screen "Filling" 800x480
   Button "Button_19" at 183,156 size 77x32; TextOff 'Aut'
      on Click: SetBit("Data_Tank1_Filling_Cmd_AutCtrl")
   TextField "Text field_26" at 286,75 size 190x23; Text 'Filling phase control'
   TextField "Text field_27" at 182,109 size 83x23; Text 'Automat'
   TextField "Text field_28" at 182,127 size 70x23; Text 'Manual'
   Button "Button_20" at 263,156 size 77x32; TextOff 'Man'
      on Click: SetBit("Data_Tank1_Filling_Cmd_ManCtrl")
   Circle "Circle_14" at 299,110 size 20x20
      Appearance <- "Data_Tank1_Filling_State_AutCtrl"
   Circle "Circle_15" at 299,130 size 20x20
      Appearance <- "Data_Tank1_Filling_State_ManCtrl"
   Button "Button_21" at 344,156 size 157x32; TextOff 'Reset done'
      on Click: SetBit("Data_Tank1_Filling_Cmd_ResetDone")
   Button "Button_22" at 183,206 size 77x32; TextOff 'Start'
      on Click: SetBit("Data_Tank1_Filling_Cmd_StartMan")
   Button "Button_23" at 263,205 size 77x32; TextOff 'Stop'
      on Click: SetBit("Data_Tank1_Filling_Cmd_StopMan")
   Button "Button_24" at 423,205 size 77x32; TextOff 'Rsume'
      on Click: SetBit("Data_Tank1_Filling_Cmd_ResumeMan")
   Button "Button_25" at 343,205 size 77x32; TextOff 'Pause'
      on Click: SetBit("Data_Tank1_Filling_Cmd_PauseMan")
   TextField "Text field_29" at 343,118 size 51x23; Text 'Done'
   Circle "Circle_16" at 460,119 size 20x20
      Appearance <- "Data_Tank1_Filling_State_Done"
   GraphicView "Graphic view_1" at 525,70 size 75x74; Picture "exit-png-cancel-cross-exit-remove-icon-512"
   Button "Button_26" at 520,72 size 76x81; TextOff 'Text'
      on Click: ActivateScreen("MainScr", 0)
   Group "Group" at 169,70 size 431x184; Picture "exit-png-cancel-cross-exit-remove-icon-512"
   SymbolLibrary "Symbol library_1" at 202,63 size 120x212
   SymbolLibrary "Symbol library_2" at 148,84 size 58x23
   SymbolLibrary "Symbol library_3" at 320,241 size 20x23
   Bar "Bar_1" at 204,63 size 117x211; MinimumValue 0; MaximumValue 2
      ProcessValue <- "Data_Tank1_WaterLevel_AIScaled"
   SymbolLibrary "Symbol library_4" at 55,31 size 94x80
      Appearance <- "Data_Tank1_ValveFill_State_StColor"
   IOField "I/O field_1" at 215,109 size 96x32; FormatPattern s9.99; Unit  m
      ProcessValue <- "Data_Tank1_WaterLevel_AIScaled"
   IOField "I/O field_2" at 216,143 size 96x32; FormatPattern 999.9; Unit  °C
      ProcessValue <- "Data_Tank1_WaterTemp_AIScaled"
   SymbolLibrary "Symbol library_6" at 226,190 size 71x61
      Appearance <- "Data_Tank1_Mixer_State_StateInt"
   Button "Button_1" at 7,233 size 77x32; TextOff 'Aut'
      on Click: SetBit("Data_Tank1_ValveFill_Cmd_AutCtrl")
   TextField "Text field_1" at 45,123 size 83x23; Text 'ValveFill'
   TextField "Text field_2" at 5,148 size 83x23; Text 'Automat'
   TextField "Text field_3" at 5,166 size 70x23; Text 'Manual'
   TextField "Text field_4" at 5,188 size 51x23; Text 'Open'
   TextField "Text field_5" at 5,206 size 65x23; Text 'Closed'
   Button "Button_2" at 86,233 size 77x32; TextOff 'Man'
      on Click: SetBit("Data_Tank1_ValveFill_Cmd_ManCtrl")
   Button "Button_3" at 7,267 size 77x32; TextOff 'Open'
      on Click: SetBit("Data_Tank1_ValveFill_Cmd_OpenMan")
   Button "Button_4" at 86,267 size 77x32; TextOff 'Close'
      on Click: SetBit("Data_Tank1_ValveFill_Cmd_CloseMan")
   Button "Button_5" at 419,209 size 77x32; TextOff 'Aut'
      on Click: SetBit("Data_Tank1_ValveDrain_Cmd_AutCtrl")
   TextField "Text field_6" at 450,99 size 104x23; Text 'ValveDrain'
   TextField "Text field_7" at 417,124 size 83x23; Text 'Automat'
   TextField "Text field_8" at 417,142 size 70x23; Text 'Manual'
   TextField "Text field_9" at 417,164 size 51x23; Text 'Open'
   TextField "Text field_10" at 417,182 size 65x23; Text 'Closed'
   Button "Button_6" at 498,209 size 77x32; TextOff 'Man'
      on Click: SetBit("Data_Tank1_Mixer_Cmd_ManCtrl")
   TextField "Text field_11" at 234,284 size 56x23; Text 'Mixer'
   TextField "Text field_12" at 185,309 size 83x23; Text 'Automat'
   TextField "Text field_13" at 185,327 size 70x23; Text 'Manual'
   TextField "Text field_14" at 185,350 size 79x23; Text 'Running'
   TextField "Text field_16" at 662,99 size 77x27; Text 'Phases'
   Button "Button_15" at 617,148 size 171x29; TextOff 'Menu filling'
      on Click: ActivateScreen("Filling", 0)
   TextField "Text field_17" at 668,124 size 61x23; Text 'Filling'
   SymbolicIOField "Symbolic I/O field_2" at 617,179 size 171x32; TextOn '1'; TextOff '0'; TextList "Phases"
      ProcessValue <- "Data_Tank1_Filling_State_Stateint"
   Button "Button_16" at 617,236 size 171x29; TextOff 'Menu draining'
      on Click: ActivateScreen("Draining", 0)
   TextField "Text field_18" at 660,213 size 82x23; Text 'Draining'
   SymbolicIOField "Symbolic I/O field_3" at 617,267 size 171x32; TextOn '1'; TextOff '0'; TextList "Phases"
      ProcessValue <- "Data_Tank1_Draining_State_StateInt"
   Button "Button_17" at 617,324 size 171x29; TextOff 'Menu mixing'
      on Click: ActivateScreen("Mixing", 0)
   TextField "Text field_19" at 669,301 size 65x23; Text 'Mixing'
   SymbolicIOField "Symbolic I/O field_4" at 617,355 size 171x32; TextOn '1'; TextOff '0'; TextList "Phases"
      ProcessValue <- "Data_Tank1_Mixing_State_StateInt"
   Button "Button_18" at 617,412 size 171x29; TextOff 'Menu heating'
      on Click: ActivateScreen("Heating", 0)
   TextField "Text field_20" at 665,390 size 76x23; Text 'Heating'
   SymbolicIOField "Symbolic I/O field_5" at 617,443 size 171x32; TextOn '1'; TextOff '0'; TextList "Phases"
      ProcessValue <- "Data_Tank1_Heating_State_StateInt"
   Button "Button_27" at 335,12 size 130x66; TextOff 'Parameters tank 1'
      on Click: ActivateScreen("Parameters", 0)
   Circle "Circle_1" at 122,149 size 20x20
      Appearance <- "Data_Tank1_ValveFill_State_AutCtrl"
   Circle "Circle_2" at 122,169 size 20x20
      Appearance <- "Data_Tank1_ValveFill_State_ManCtrl"
   Circle "Circle_3" at 122,189 size 20x20
      Appearance <- "Data_Tank1_ValveFill_State_Open"
   Circle "Circle_4" at 122,209 size 20x20
      Appearance <- "Data_Tank1_ValveFill_State_Closed"
   Circle "Circle_5" at 534,125 size 20x20
      Appearance <- "Data_Tank1_ValveDrain_State_AutCtrl"
   Circle "Circle_6" at 534,145 size 20x20
      Appearance <- "Data_Tank1_ValveDrain_State_ManCtrl"
   Circle "Circle_7" at 534,165 size 20x20
      Appearance <- "Data_Tank1_ValveDrain_State_Open"
   Circle "Circle_8" at 534,185 size 20x20
      Appearance <- "Data_Tank1_ValveDrain_State_Closed"
   TextField "Text field_21" at 427,285 size 156x23; Text 'Heating element'
   TextField "Text field_22" at 418,310 size 83x23; Text 'Automat'
   TextField "Text field_23" at 418,328 size 70x23; Text 'Manual'
   TextField "Text field_24" at 422,350 size 157x23; Text 'Manual heat pwr'

screen "Draining" 800x480
   TextField "Text field_26" at 286,163 size 211x23; Text 'Draining phase control'
   TextField "Text field_27" at 182,197 size 83x23; Text 'Automat'
   TextField "Text field_28" at 182,215 size 70x23; Text 'Manual'
   TextField "Text field_29" at 343,206 size 51x23; Text 'Done'
   GraphicView "Graphic view_1" at 525,158 size 75x74; Picture "exit-png-cancel-cross-exit-remove-icon-512"
   Button "Button_26" at 520,160 size 76x81; TextOff 'Text'
      on Click: ActivateScreen("MainScr", 0)
   Circle "Circle_5" at 288,199 size 20x20
      Appearance <- "Data_Tank1_Draining_State_AutCtrl"
   Circle "Circle_6" at 288,220 size 20x20
      Appearance <- "Data_Tank1_Draining_State_ManCtrl"
   Circle "Circle_10" at 440,201 size 35x35
      Appearance <- "Data_Tank1_Draining_State_Done"
   Button "Button_9" at 183,251 size 77x32; TextOff 'Aut'
      on Click: SetBit("Data_Tank1_Draining_Cmd_AutCtrl")
   Button "Button_10" at 258,251 size 77x32; TextOff 'Man'
      on Click: SetBit("Data_Tank1_Draining_Cmd_ManCtrl")
   Button "Button_11" at 344,252 size 158x32; TextOff 'Reset Done'
      on Click: SetBit("Data_Tank1_Draining_Cmd_ResetDone")
   Button "Button_12" at 183,285 size 77x32; TextOff 'Start'
      on Click: SetBit("Data_Tank1_Draining_Cmd_StartMan")
   Button "Button_13" at 258,285 size 77x32; TextOff 'Stop'
      on Click: SetBit("Data_Tank1_Draining_Cmd_StopMan")
   Button "Button_14" at 345,286 size 77x32; TextOff 'Pause'
      on Click: SetBit("Data_Tank1_Draining_Cmd_PauseMan")
   Button "Button_19" at 422,286 size 77x32; TextOff 'Rsume'
      on Click: SetBit("Data_Tank1_Draining_Cmd_ResumeMan")
   SymbolLibrary "Symbol library_1" at 202,63 size 120x212
   SymbolLibrary "Symbol library_2" at 148,84 size 58x23
   SymbolLibrary "Symbol library_3" at 320,241 size 20x23
   Bar "Bar_1" at 204,63 size 117x211; MinimumValue 0; MaximumValue 2
      ProcessValue <- "Data_Tank1_WaterLevel_AIScaled"
   SymbolLibrary "Symbol library_4" at 55,31 size 94x80
      Appearance <- "Data_Tank1_ValveFill_State_StColor"
   SymbolLibrary "Symbol library_5" at 314,188 size 94x80
      Appearance <- "Data_Tank1_ValveDrain_State_StColor"
   IOField "I/O field_1" at 215,109 size 96x32; FormatPattern s9.99; Unit  m
      ProcessValue <- "Data_Tank1_WaterLevel_AIScaled"
   IOField "I/O field_2" at 216,143 size 96x32; FormatPattern 999.9; Unit  °C
      ProcessValue <- "Data_Tank1_WaterTemp_AIScaled"
   SymbolLibrary "Symbol library_6" at 226,190 size 71x61
      Appearance <- "Data_Tank1_Mixer_State_StateInt"
   Button "Button_1" at 7,233 size 77x32; TextOff 'Aut'
      on Click: SetBit("Data_Tank1_ValveFill_Cmd_AutCtrl")
   TextField "Text field_1" at 45,123 size 83x23; Text 'ValveFill'
   TextField "Text field_2" at 5,148 size 83x23; Text 'Automat'
   TextField "Text field_3" at 5,166 size 70x23; Text 'Manual'
   TextField "Text field_4" at 5,188 size 51x23; Text 'Open'
   TextField "Text field_5" at 5,206 size 65x23; Text 'Closed'
   Button "Button_2" at 86,233 size 77x32; TextOff 'Man'
      on Click: SetBit("Data_Tank1_ValveFill_Cmd_ManCtrl")
   Button "Button_3" at 7,267 size 77x32; TextOff 'Open'
      on Click: SetBit("Data_Tank1_ValveFill_Cmd_OpenMan")
   Button "Button_4" at 86,267 size 77x32; TextOff 'Close'
      on Click: SetBit("Data_Tank1_ValveFill_Cmd_CloseMan")
   Button "Button_5" at 419,209 size 77x32; TextOff 'Aut'
      on Click: SetBit("Data_Tank1_ValveDrain_Cmd_AutCtrl")
   TextField "Text field_6" at 450,99 size 104x23; Text 'ValveDrain'
   TextField "Text field_7" at 417,124 size 83x23; Text 'Automat'
   TextField "Text field_8" at 417,142 size 70x23; Text 'Manual'
   TextField "Text field_9" at 417,164 size 51x23; Text 'Open'
   TextField "Text field_10" at 417,182 size 65x23; Text 'Closed'
   Button "Button_6" at 498,209 size 77x32; TextOff 'Man'
      on Click: SetBit("Data_Tank1_Mixer_Cmd_ManCtrl")
   Button "Button_7" at 419,243 size 77x32; TextOff 'Open'
      on Click: SetBit("Data_Tank1_ValveDrain_Cmd_OpenMan")
   Button "Button_8" at 498,243 size 77x32; TextOff 'Close'
      on Click: SetBit("Data_Tank1_ValveDrain_Cmd_CloseMan")
   TextField "Text field_11" at 234,284 size 56x23; Text 'Mixer'
   TextField "Text field_12" at 185,309 size 83x23; Text 'Automat'
   TextField "Text field_13" at 185,327 size 70x23; Text 'Manual'
   TextField "Text field_14" at 185,350 size 79x23; Text 'Running'
   TextField "Text field_16" at 662,99 size 77x27; Text 'Phases'
   Button "Button_15" at 617,148 size 171x29; TextOff 'Menu filling'
      on Click: ActivateScreen("Filling", 0)
   TextField "Text field_17" at 668,124 size 61x23; Text 'Filling'
   SymbolicIOField "Symbolic I/O field_2" at 617,179 size 171x32; TextOn '1'; TextOff '0'; TextList "Phases"
      ProcessValue <- "Data_Tank1_Filling_State_Stateint"
   Button "Button_16" at 617,236 size 171x29; TextOff 'Menu draining'
      on Click: ActivateScreen("Draining", 0)
   TextField "Text field_18" at 660,213 size 82x23; Text 'Draining'
   SymbolicIOField "Symbolic I/O field_3" at 617,267 size 171x32; TextOn '1'; TextOff '0'; TextList "Phases"
      ProcessValue <- "Data_Tank1_Draining_State_StateInt"
   Button "Button_17" at 617,324 size 171x29; TextOff 'Menu mixing'
      on Click: ActivateScreen("Mixing", 0)
   TextField "Text field_19" at 669,301 size 65x23; Text 'Mixing'
   SymbolicIOField "Symbolic I/O field_4" at 617,355 size 171x32; TextOn '1'; TextOff '0'; TextList "Phases"
      ProcessValue <- "Data_Tank1_Mixing_State_StateInt"
   Button "Button_18" at 617,412 size 171x29; TextOff 'Menu heating'
      on Click: ActivateScreen("Heating", 0)
   TextField "Text field_20" at 665,390 size 76x23; Text 'Heating'
   SymbolicIOField "Symbolic I/O field_5" at 617,443 size 171x32; TextOn '1'; TextOff '0'; TextList "Phases"
      ProcessValue <- "Data_Tank1_Heating_State_StateInt"
   TextField "Text field_21" at 427,291 size 156x23; Text 'Heating element'
   TextField "Text field_22" at 418,316 size 83x23; Text 'Automat'
   Button "Button_27" at 335,12 size 130x66; TextOff 'Parameters tank 1'
      on Click: ActivateScreen("Parameters", 0)
   Circle "Circle_1" at 122,149 size 20x20
      Appearance <- "Data_Tank1_ValveFill_State_AutCtrl"
   Circle "Circle_2" at 122,169 size 20x20
      Appearance <- "Data_Tank1_ValveFill_State_ManCtrl"
   Circle "Circle_3" at 122,189 size 20x20
      Appearance <- "Data_Tank1_ValveFill_State_Open"
   Circle "Circle_4" at 122,209 size 20x20
      Appearance <- "Data_Tank1_ValveFill_State_Closed"
   Circle "Circle_7" at 534,165 size 20x20
      Appearance <- "Data_Tank1_ValveDrain_State_Open"
   Circle "Circle_8" at 534,185 size 20x20
      Appearance <- "Data_Tank1_ValveDrain_State_Closed"
   Circle "Circle_9" at 302,310 size 20x20
      Appearance <- "Data_Tank1_Mixer_State_AutCtrl"
   Circle "Circle_11" at 535,317 size 20x20
      Appearance <- "Data_Tank1_Heating_Cmd_AutCtrl"
   Circle "Circle_13" at 535,317 size 20x20
      Appearance <- "Data_Tank1_Heating_State_AutCtrl"
   TextField "Text field_23" at 427,285 size 156x23; Text 'Heating element'
   TextField "Text field_24" at 418,310 size 83x23; Text 'Automat'
   TextField "Text field_25" at 418,328 size 70x23; Text 'Manual'
   TextField "Text field_30" at 422,350 size 157x23; Text 'Manual heat pwr'
   Circle "Circle_17" at 535,311 size 20x20
      Appearance <- "Data_Tank1_Heater_State_AutCtrl"

screen "Parameters" 800x480
   Button "Button_19" at 659,404 size 130x66; TextOff 'Main screen'
      on Click: ActivateScreen("MainScr", 0)
   TextField "Text field_24" at 62,105 size 97x23; Text 'Level max'
   IOField "I/O field_3" at 60,140 size 96x32; FormatPattern 9.99; Unit  m
      ProcessValue <- "Data_Tank1_Filling_Param_FillLevel"
   TextField "Text field_1" at 67,203 size 92x23; Text 'Level min'
   IOField "I/O field_1" at 58,230 size 96x32; FormatPattern 9.99; Unit  m
      ProcessValue <- "Data_Tank1_Draining_Param_DrainLevel"
   TextField "Text field_2" at 243,102 size 123x23; Text 'Temperature'
   IOField "I/O field_2" at 252,134 size 96x32; FormatPattern 99.9; Unit  °C
      ProcessValue <- "Data_Tank1_Heating_Param_ReqTemp"
   TextField "Text field_4" at 447,103 size 112x23; Text 'Mixing time'
   IOField "I/O field_4" at 451,131 size 96x32; FormatPattern 99; Unit  s
      ProcessValue <- "Data_Tank1_Mixing_Param_TimeSec"
   Bar "Bar_1" at 239,196 size 128x230; MinimumValue 0; MaximumValue 100
      ProcessValue <- "Data_Tank1_Heating_Param_ReqTemp"
*)